(* Logix 5000 project; controller PLC_MCC1201_220AP1 vendor 1 type 14 code 164 rev 35.11; software revision 35.00; part 11 of 25 *)
(* tags used below, declared in another part *)
   AFI : ALIAS FOR B3[7].15;
   B175 : DINT[1];
   B176 : DINT[1];
   B180 : DINT[10];
   BT181_000 : MESSAGE;
   BT181_004 : MESSAGE;
   BT181_005 : MESSAGE;
   BT181_006 : MESSAGE;
   BT181_007 : MESSAGE;
   BT181_008 : MESSAGE;
   C183 : COUNTER[3];
   ConsumedFromCullet : UDT_CONSUMED_CULLET;
   ConsumedFromMCC1300 : UDT_CONSUMED_NEXT;
   CPU_FaultRecord : SYS_FaultRecord;
   CPU_LastFaultRecord : SYS_FaultRecord;
   From_Cullet : DINT[10];
   HMI_Always_ON : BOOL;   // HMI Always ON
   I : INT[128];
   M202_M1_DR : AXIS_CIP_DRIVE;
   M202_M1_DR_IN_MAJ : MOTION_INSTRUCTION;
   M202_M1_DR_IN_MAM : MOTION_INSTRUCTION;
   M202_M1_DR_IN_MAR : MOTION_INSTRUCTION;
   M202_M1_DR_IN_MAS : MOTION_INSTRUCTION;
   M202_M1_DR_IN_MCD : MOTION_INSTRUCTION;
   M202_M1_DR_IN_MRP : MOTION_INSTRUCTION;
   M202_M1_DR_OUT_MAJ : MOTION_INSTRUCTION;
   M202_M1_DR_OUT_MAM : MOTION_INSTRUCTION;
   M202_M1_DR_OUT_MAR : MOTION_INSTRUCTION;
   M202_M1_DR_OUT_MAS : MOTION_INSTRUCTION;
   M202_M1_DR_OUT_MCD : MOTION_INSTRUCTION;
   M202_M1_DR_OUT_MRP : MOTION_INSTRUCTION;
   M203_M1_DR : AXIS_CIP_DRIVE;
   M203_M1_DR_IN_MAJ : MOTION_INSTRUCTION;
   M203_M1_DR_IN_MAM : MOTION_INSTRUCTION;
   M203_M1_DR_IN_MAR : MOTION_INSTRUCTION;
   M203_M1_DR_IN_MAS : MOTION_INSTRUCTION;
   M203_M1_DR_IN_MCD : MOTION_INSTRUCTION;
   M203_M1_DR_IN_MRP : MOTION_INSTRUCTION;
   M203_M1_DR_OUT_MAJ : MOTION_INSTRUCTION;
   M203_M1_DR_OUT_MAM : MOTION_INSTRUCTION;
   M203_M1_DR_OUT_MAR : MOTION_INSTRUCTION;
   M203_M1_DR_OUT_MAS : MOTION_INSTRUCTION;
   M203_M1_DR_OUT_MCD : MOTION_INSTRUCTION;
   M203_M1_DR_OUT_MRP : MOTION_INSTRUCTION;
   M203DROP : MAC_DROPCONV;
   M204_M1_DR : AXIS_CIP_DRIVE;
   M204_M1_DR_IN_MAJ : MOTION_INSTRUCTION;
   M204_M1_DR_IN_MAM : MOTION_INSTRUCTION;
   M204_M1_DR_IN_MAR : MOTION_INSTRUCTION;
   M204_M1_DR_IN_MAS : MOTION_INSTRUCTION;
   M204_M1_DR_IN_MCD : MOTION_INSTRUCTION;
   M204_M1_DR_IN_MRP : MOTION_INSTRUCTION;
   M204_M1_DR_OUT_MAJ : MOTION_INSTRUCTION;
   M204_M1_DR_OUT_MAM : MOTION_INSTRUCTION;
   M204_M1_DR_OUT_MAR : MOTION_INSTRUCTION;
   M204_M1_DR_OUT_MAS : MOTION_INSTRUCTION;
   M204_M1_DR_OUT_MCD : MOTION_INSTRUCTION;
   M204_M1_DR_OUT_MRP : MOTION_INSTRUCTION;
   M205BREAKER : MAC_BREAKER;
   M206_M1_DR : AXIS_CIP_DRIVE;
   M206_M1_DR_IN_MAJ : MOTION_INSTRUCTION;
   M206_M1_DR_IN_MAM : MOTION_INSTRUCTION;
   M206_M1_DR_IN_MAR : MOTION_INSTRUCTION;
   M206_M1_DR_IN_MAS : MOTION_INSTRUCTION;
   M206_M1_DR_IN_MCD : MOTION_INSTRUCTION;
   M206_M1_DR_IN_MRP : MOTION_INSTRUCTION;
   M206_M1_DR_OUT_MAJ : MOTION_INSTRUCTION;
   M206_M1_DR_OUT_MAM : MOTION_INSTRUCTION;
   M206_M1_DR_OUT_MAR : MOTION_INSTRUCTION;
   M206_M1_DR_OUT_MAS : MOTION_INSTRUCTION;
   M206_M1_DR_OUT_MCD : MOTION_INSTRUCTION;
   M206_M1_DR_OUT_MRP : MOTION_INSTRUCTION;
   M207_M1_DR : AXIS_CIP_DRIVE;
   M207_M1_DR_IN_MAJ : MOTION_INSTRUCTION;
   M207_M1_DR_IN_MAM : MOTION_INSTRUCTION;
   M207_M1_DR_IN_MAR : MOTION_INSTRUCTION;
   M207_M1_DR_IN_MAS : MOTION_INSTRUCTION;
   M207_M1_DR_IN_MCD : MOTION_INSTRUCTION;
   M207_M1_DR_IN_MRP : MOTION_INSTRUCTION;
   M207_M1_DR_OUT_MAJ : MOTION_INSTRUCTION;
   M207_M1_DR_OUT_MAM : MOTION_INSTRUCTION;
   M207_M1_DR_OUT_MAR : MOTION_INSTRUCTION;
   M207_M1_DR_OUT_MAS : MOTION_INSTRUCTION;
   M207_M1_DR_OUT_MCD : MOTION_INSTRUCTION;
   M207_M1_DR_OUT_MRP : MOTION_INSTRUCTION;
   M208_M1_DR : AXIS_CIP_DRIVE;
   M208_M1_DR_IN_MAJ : MOTION_INSTRUCTION;
   M208_M1_DR_IN_MAM : MOTION_INSTRUCTION;
   M208_M1_DR_IN_MAR : MOTION_INSTRUCTION;
   M208_M1_DR_IN_MAS : MOTION_INSTRUCTION;
   M208_M1_DR_IN_MCD : MOTION_INSTRUCTION;
   M208_M1_DR_IN_MRP : MOTION_INSTRUCTION;
   M208_M1_DR_OUT_MAJ : MOTION_INSTRUCTION;
   M208_M1_DR_OUT_MAM : MOTION_INSTRUCTION;
   M208_M1_DR_OUT_MAR : MOTION_INSTRUCTION;
   M208_M1_DR_OUT_MAS : MOTION_INSTRUCTION;
   M208_M1_DR_OUT_MCD : MOTION_INSTRUCTION;
   M208_M1_DR_OUT_MRP : MOTION_INSTRUCTION;
   M209_M1_DR : AXIS_CIP_DRIVE;
   M209_M1_DR_IN_MAJ : MOTION_INSTRUCTION;
   M209_M1_DR_IN_MAM : MOTION_INSTRUCTION;
   M209_M1_DR_IN_MAR : MOTION_INSTRUCTION;
   M209_M1_DR_IN_MAS : MOTION_INSTRUCTION;
   M209_M1_DR_IN_MCD : MOTION_INSTRUCTION;
   M209_M1_DR_IN_MRP : MOTION_INSTRUCTION;
   M209_M1_DR_OUT_MAJ : MOTION_INSTRUCTION;
   M209_M1_DR_OUT_MAM : MOTION_INSTRUCTION;
   M209_M1_DR_OUT_MAR : MOTION_INSTRUCTION;
   M209_M1_DR_OUT_MAS : MOTION_INSTRUCTION;
   M209_M1_DR_OUT_MCD : MOTION_INSTRUCTION;
   M209_M1_DR_OUT_MRP : MOTION_INSTRUCTION;
   M210_M1_DR : AXIS_CIP_DRIVE;
   M210_M1_DR_IN_MAJ : MOTION_INSTRUCTION;
   M210_M1_DR_IN_MAM : MOTION_INSTRUCTION;
   M210_M1_DR_IN_MAR : MOTION_INSTRUCTION;
   M210_M1_DR_IN_MAS : MOTION_INSTRUCTION;
   M210_M1_DR_IN_MCD : MOTION_INSTRUCTION;
   M210_M1_DR_IN_MRP : MOTION_INSTRUCTION;
   M210_M1_DR_OUT_MAJ : MOTION_INSTRUCTION;
   M210_M1_DR_OUT_MAM : MOTION_INSTRUCTION;
   M210_M1_DR_OUT_MAR : MOTION_INSTRUCTION;
   M210_M1_DR_OUT_MAS : MOTION_INSTRUCTION;
   M210_M1_DR_OUT_MCD : MOTION_INSTRUCTION;
   M210_M1_DR_OUT_MRP : MOTION_INSTRUCTION;
   M211_M1_DR : AXIS_CIP_DRIVE;
   M211_M1_DR_IN_MAJ : MOTION_INSTRUCTION;
   M211_M1_DR_IN_MAM : MOTION_INSTRUCTION;
   M211_M1_DR_IN_MAR : MOTION_INSTRUCTION;
   M211_M1_DR_IN_MAS : MOTION_INSTRUCTION;
   M211_M1_DR_IN_MCD : MOTION_INSTRUCTION;
   M211_M1_DR_IN_MRP : MOTION_INSTRUCTION;
   M211_M1_DR_OUT_MAJ : MOTION_INSTRUCTION;
   M211_M1_DR_OUT_MAM : MOTION_INSTRUCTION;
   M211_M1_DR_OUT_MAR : MOTION_INSTRUCTION;
   M211_M1_DR_OUT_MAS : MOTION_INSTRUCTION;
   M211_M1_DR_OUT_MCD : MOTION_INSTRUCTION;
   M211_M1_DR_OUT_MRP : MOTION_INSTRUCTION;
   M212_M1_DR : AXIS_CIP_DRIVE;
   M212_M1_DR_IN_MAJ : MOTION_INSTRUCTION;
   M212_M1_DR_IN_MAM : MOTION_INSTRUCTION;
   M212_M1_DR_IN_MAR : MOTION_INSTRUCTION;
   M212_M1_DR_IN_MAS : MOTION_INSTRUCTION;
   M212_M1_DR_IN_MCD : MOTION_INSTRUCTION;
   M212_M1_DR_IN_MRP : MOTION_INSTRUCTION;
   M212_M1_DR_OUT_MAJ : MOTION_INSTRUCTION;
   M212_M1_DR_OUT_MAM : MOTION_INSTRUCTION;
   M212_M1_DR_OUT_MAR : MOTION_INSTRUCTION;
   M212_M1_DR_OUT_MAS : MOTION_INSTRUCTION;
   M212_M1_DR_OUT_MCD : MOTION_INSTRUCTION;
   M212_M1_DR_OUT_MRP : MOTION_INSTRUCTION;
   M213_M1_DR : AXIS_CIP_DRIVE;
   M213_M1_DR_IN_MAJ : MOTION_INSTRUCTION;
   M213_M1_DR_IN_MAM : MOTION_INSTRUCTION;
   M213_M1_DR_IN_MAR : MOTION_INSTRUCTION;
   M213_M1_DR_IN_MAS : MOTION_INSTRUCTION;
   M213_M1_DR_IN_MCD : MOTION_INSTRUCTION;
   M213_M1_DR_IN_MRP : MOTION_INSTRUCTION;
   M213_M1_DR_OUT_MAJ : MOTION_INSTRUCTION;
   M213_M1_DR_OUT_MAM : MOTION_INSTRUCTION;
   M213_M1_DR_OUT_MAR : MOTION_INSTRUCTION;
   M213_M1_DR_OUT_MAS : MOTION_INSTRUCTION;
   M213_M1_DR_OUT_MCD : MOTION_INSTRUCTION;
   M213_M1_DR_OUT_MRP : MOTION_INSTRUCTION;
   M213A_M1_DR_IN_MAJ : MOTION_INSTRUCTION;
   M213A_M1_DR_IN_MAM : MOTION_INSTRUCTION;
   M213A_M1_DR_IN_MAR : MOTION_INSTRUCTION;
   M213A_M1_DR_IN_MAS : MOTION_INSTRUCTION;
   M213A_M1_DR_IN_MCD : MOTION_INSTRUCTION;
   M213A_M1_DR_IN_MRP : MOTION_INSTRUCTION;
   M213A_M1_DR_OUT_MAJ : MOTION_INSTRUCTION;
   M213A_M1_DR_OUT_MAM : MOTION_INSTRUCTION;
   M213A_M1_DR_OUT_MAR : MOTION_INSTRUCTION;
   M213A_M1_DR_OUT_MAS : MOTION_INSTRUCTION;
   M213A_M1_DR_OUT_MCD : MOTION_INSTRUCTION;
   M213A_M1_DR_OUT_MRP : MOTION_INSTRUCTION;
   M213B_M1_DR_IN_MAJ : MOTION_INSTRUCTION;
   M213B_M1_DR_IN_MAM : MOTION_INSTRUCTION;
   M213B_M1_DR_IN_MAR : MOTION_INSTRUCTION;
   M213B_M1_DR_IN_MAS : MOTION_INSTRUCTION;
   M213B_M1_DR_IN_MCD : MOTION_INSTRUCTION;
   M213B_M1_DR_IN_MRP : MOTION_INSTRUCTION;
   M213B_M1_DR_OUT_MAJ : MOTION_INSTRUCTION;
   M213B_M1_DR_OUT_MAM : MOTION_INSTRUCTION;
   M213B_M1_DR_OUT_MAR : MOTION_INSTRUCTION;
   M213B_M1_DR_OUT_MAS : MOTION_INSTRUCTION;
   M213B_M1_DR_OUT_MCD : MOTION_INSTRUCTION;
   M213B_M1_DR_OUT_MRP : MOTION_INSTRUCTION;
   M214_M1_DR : AXIS_CIP_DRIVE;
   M214_M1_DR_IN_MAJ : MOTION_INSTRUCTION;
   M214_M1_DR_IN_MAM : MOTION_INSTRUCTION;
   M214_M1_DR_IN_MAR : MOTION_INSTRUCTION;
   M214_M1_DR_IN_MAS : MOTION_INSTRUCTION;
   M214_M1_DR_IN_MCD : MOTION_INSTRUCTION;
   M214_M1_DR_IN_MRP : MOTION_INSTRUCTION;
   M214_M1_DR_OUT_MAJ : MOTION_INSTRUCTION;
   M214_M1_DR_OUT_MAM : MOTION_INSTRUCTION;
   M214_M1_DR_OUT_MAR : MOTION_INSTRUCTION;
   M214_M1_DR_OUT_MAS : MOTION_INSTRUCTION;
   M214_M1_DR_OUT_MCD : MOTION_INSTRUCTION;
   M214_M1_DR_OUT_MRP : MOTION_INSTRUCTION;
   M215_M1_DR : AXIS_CIP_DRIVE;
   M215_M1_DR_IN_MAJ : MOTION_INSTRUCTION;
   M215_M1_DR_IN_MAM : MOTION_INSTRUCTION;
   M215_M1_DR_IN_MAR : MOTION_INSTRUCTION;
   M215_M1_DR_IN_MAS : MOTION_INSTRUCTION;
   M215_M1_DR_IN_MCD : MOTION_INSTRUCTION;
   M215_M1_DR_IN_MRP : MOTION_INSTRUCTION;
   M215_M1_DR_OUT_MAJ : MOTION_INSTRUCTION;
   M215_M1_DR_OUT_MAM : MOTION_INSTRUCTION;
   M215_M1_DR_OUT_MAR : MOTION_INSTRUCTION;
   M215_M1_DR_OUT_MAS : MOTION_INSTRUCTION;
   M215_M1_DR_OUT_MCD : MOTION_INSTRUCTION;
   M215_M1_DR_OUT_MRP : MOTION_INSTRUCTION;
   M216_M1_DR : AXIS_CIP_DRIVE;
   M216_M1_DR_IN_MAJ : MOTION_INSTRUCTION;
   M216_M1_DR_IN_MAM : MOTION_INSTRUCTION;
   M216_M1_DR_IN_MAR : MOTION_INSTRUCTION;
   M216_M1_DR_IN_MAS : MOTION_INSTRUCTION;
   M216_M1_DR_IN_MCD : MOTION_INSTRUCTION;
   M216_M1_DR_IN_MRP : MOTION_INSTRUCTION;
   M216_M1_DR_OUT_MAJ : MOTION_INSTRUCTION;
   M216_M1_DR_OUT_MAM : MOTION_INSTRUCTION;
   M216_M1_DR_OUT_MAR : MOTION_INSTRUCTION;
   M216_M1_DR_OUT_MAS : MOTION_INSTRUCTION;
   M216_M1_DR_OUT_MCD : MOTION_INSTRUCTION;
   M216_M1_DR_OUT_MRP : MOTION_INSTRUCTION;
   M217_M1_DR : AXIS_CIP_DRIVE;
   M217_M1_DR_IN_MAJ : MOTION_INSTRUCTION;
   M217_M1_DR_IN_MAM : MOTION_INSTRUCTION;
   M217_M1_DR_IN_MAR : MOTION_INSTRUCTION;
   M217_M1_DR_IN_MAS : MOTION_INSTRUCTION;
   M217_M1_DR_IN_MCD : MOTION_INSTRUCTION;
   M217_M1_DR_IN_MRP : MOTION_INSTRUCTION;
   M217_M1_DR_OUT_MAJ : MOTION_INSTRUCTION;
   M217_M1_DR_OUT_MAM : MOTION_INSTRUCTION;
   M217_M1_DR_OUT_MAR : MOTION_INSTRUCTION;
   M217_M1_DR_OUT_MAS : MOTION_INSTRUCTION;
   M217_M1_DR_OUT_MCD : MOTION_INSTRUCTION;
   M217_M1_DR_OUT_MRP : MOTION_INSTRUCTION;
   M218_M1_DR : AXIS_CIP_DRIVE;
   M218_M1_DR_IN_MAJ : MOTION_INSTRUCTION;
   M218_M1_DR_IN_MAM : MOTION_INSTRUCTION;
   M218_M1_DR_IN_MAR : MOTION_INSTRUCTION;
   M218_M1_DR_IN_MAS : MOTION_INSTRUCTION;
   M218_M1_DR_IN_MCD : MOTION_INSTRUCTION;
   M218_M1_DR_IN_MRP : MOTION_INSTRUCTION;
   M218_M1_DR_OUT_MAJ : MOTION_INSTRUCTION;
   M218_M1_DR_OUT_MAM : MOTION_INSTRUCTION;
   M218_M1_DR_OUT_MAR : MOTION_INSTRUCTION;
   M218_M1_DR_OUT_MAS : MOTION_INSTRUCTION;
(* CommandLogic, continued *)

ROUTINE Main   (* ladder *)
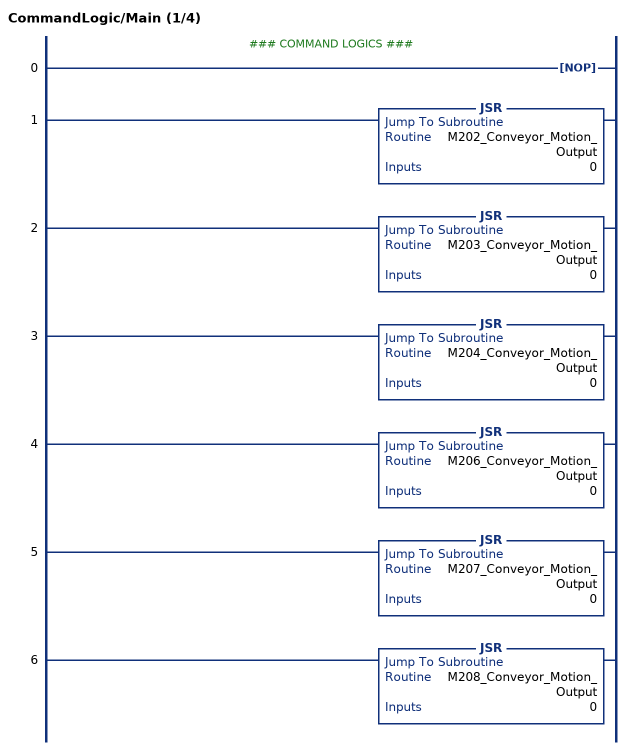
   // ### COMMAND LOGICS ###
   0: NOP();
   1: JSR(M202_Conveyor_Motion_Output,0);
   2: JSR(M203_Conveyor_Motion_Output,0);
   3: JSR(M204_Conveyor_Motion_Output,0);
   4: JSR(M206_Conveyor_Motion_Output,0);
   5: JSR(M207_Conveyor_Motion_Output,0);
   6: JSR(M208_Conveyor_Motion_Output,0);
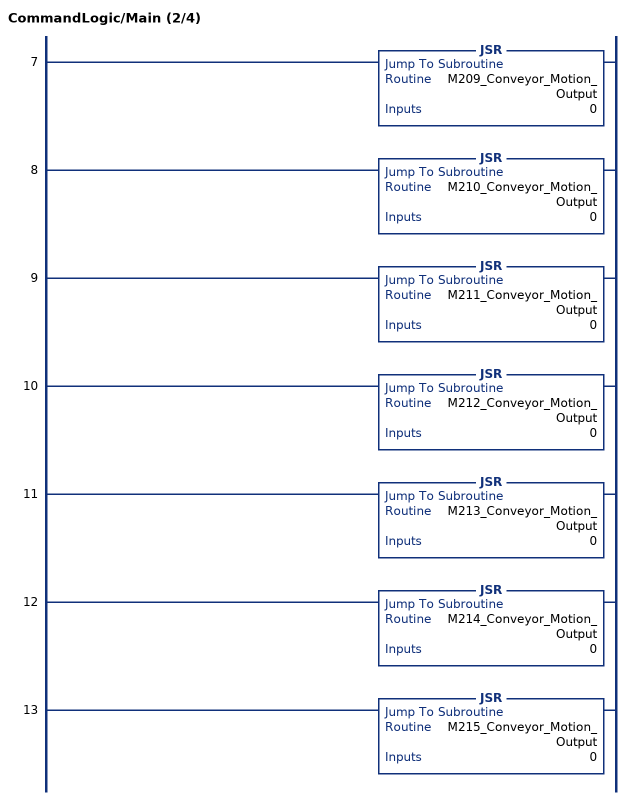
   7: JSR(M209_Conveyor_Motion_Output,0);
   8: JSR(M210_Conveyor_Motion_Output,0);
   9: JSR(M211_Conveyor_Motion_Output,0);
   10: JSR(M212_Conveyor_Motion_Output,0);
   11: JSR(M213_Conveyor_Motion_Output,0);
   12: JSR(M214_Conveyor_Motion_Output,0);
   13: JSR(M215_Conveyor_Motion_Output,0);
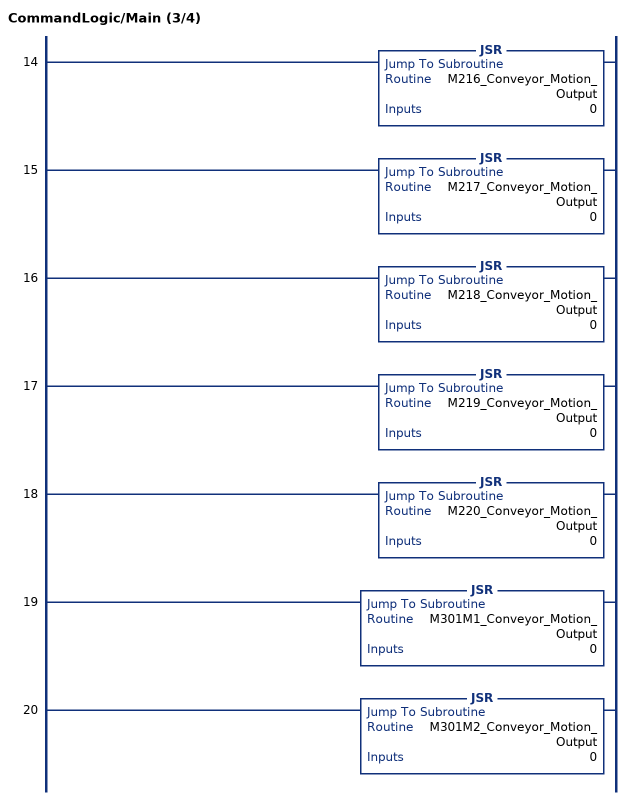
   14: JSR(M216_Conveyor_Motion_Output,0);
   15: JSR(M217_Conveyor_Motion_Output,0);
   16: JSR(M218_Conveyor_Motion_Output,0);
   17: JSR(M219_Conveyor_Motion_Output,0);
   18: JSR(M220_Conveyor_Motion_Output,0);
   19: JSR(M301M1_Conveyor_Motion_Output,0);
   20: JSR(M301M2_Conveyor_Motion_Output,0);
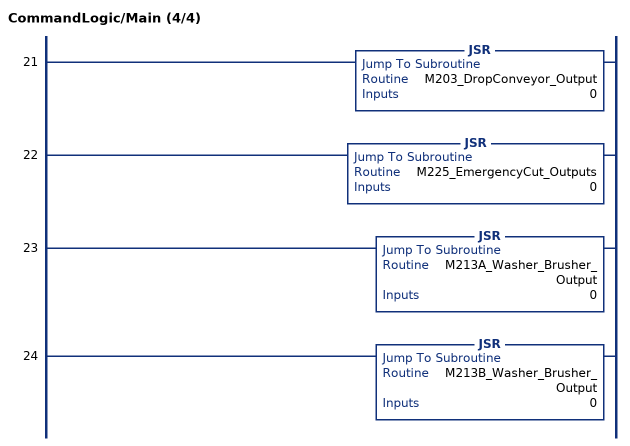
   21: JSR(M203_DropConveyor_Output,0);
   22: JSR(M225_EmergencyCut_Outputs,0);
   23: JSR(M213A_Washer_Brusher_Output,0);
   24: JSR(M213B_Washer_Brusher_Output,0);
END_ROUTINE
END_PROGRAM

PROGRAM ControllerErrors   (* main routine Main *)

ROUTINE Main   (* ladder *)
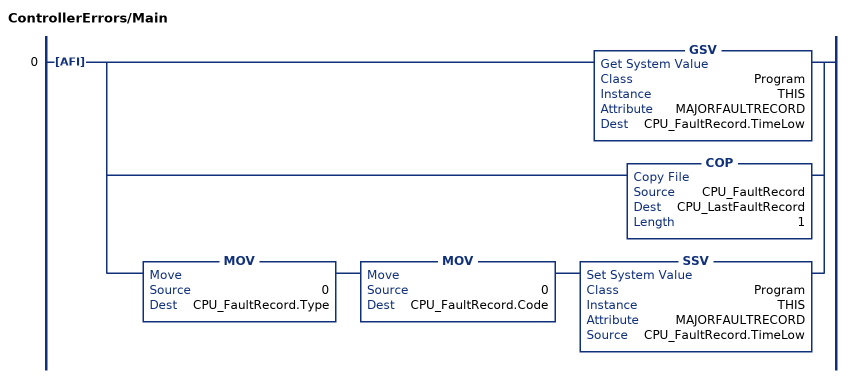
   0: AFI()[GSV(Program,THIS,MAJORFAULTRECORD,CPU_FaultRecord.TimeLow) ,COP(CPU_FaultRecord,CPU_LastFaultRecord,1) ,MOV(0,CPU_FaultRecord.Type) MOV(0,CPU_FaultRecord.Code) SSV(Program,THIS,MAJORFAULTRECORD,CPU_FaultRecord.TimeLow) ];
END_ROUTINE
END_PROGRAM

PROGRAM MainProgram   (* main routine MainRoutine *)
VAR
   dMaxLehrSpeed : DINT := 20000;
   dMinLehrSpeed : DINT := 1270;
   GP_M225_AccessArea_FarSide : GP_AccessArea := (IN_xConditionOkForcedAccess := 1);
   GP_M225_AccessArea_FarSide_STC : GP_AccessArea_STC := (OSR_xAccessRequest := 1, OSR_xAccessAcceptedAndButtonReleased := 1, OSR_xRemoveAccess := 1, OSR_xRemoveAccessNotAccepted := 1);
   GP_M225_AccessArea_OpSide : GP_AccessArea := (IN_xConditionOkForcedAccess := 1);
   GP_M225_AccessArea_OpSide_STC : GP_AccessArea_STC := (OSR_xAccessRequest := 1, OSR_xAccessAcceptedAndButtonReleased := 1, OSR_xRemoveAccess := 1, OSR_xRemoveAccessNotAccepted := 1);
   GP_RibbonTracking_GetRibbonData : GP_RibbonTracking_GetRibbonData;
   GP_RibbonTracking_UpdateGlassBreak : GP_RibbonTracking_UpdateGlassBreak;
   LEHR_dActualSpeedValue_mm_min : DINT;
   LEHR_dActualSpeedValueToConveyor_mm_min : DINT;
   LEHR_dLehrPositionAdvancement : DINT;
   SnaprollHMW_dOffset_cmm : DINT;
   SnaprollUPS_DistanceFromSnaproll_cmm : DINT := 4663000;
   SnaprollUPS_xOS_NewCut : BOOL;
   SnaprollUPS_xOSR : BOOL;
   SnaprollUPS_xOutputRise : BOOL;
   tmOF_retainSnaprolUPS : TIMER;
   TMP_dDistanceBetweenCut : DINT := 273986272;
   TMP_dDummy : DINT := 4215000;
   TMP_dEncoderCutPosition : DINT;
   TMP_dSnaprollCut_cmm : DINT := 4663000;
   TMP_dValue : DINT;
   TMP_xCutOnSnaproll_cmm : BOOL;
   TMP_xDummy : BOOL;
   TMP_xSimulationMode : BOOL;
   xAlwaysOFF : BOOL;
   xAlwaysON : BOOL := 1;
   xDebugOFF : BOOL;
END_VAR

ROUTINE _010_Input_Mapping   (* structured text *)
   
   //Always ON bit for HMI
   HMI_Always_ON := 1;
   
   //INPUT
   
   //Z200 UPS ZONE (UNTIL MAIN CRUSHER)
   Z200_UPS.INPUT_x24vdcVoltageOn := A152AP1:1:I.Pt00.Data;
   Z200_UPS.INPUT_xUPSEmergencyON := A152AP1:1:I.Pt04.Data;
   Z200_UPS.INPUT_xEmLocUps1 := A152AP1:6:I.Pt11.Data; //A33SB2 UPS Emergency Button M203DROP OPERATOR SIDE
   Z200_UPS.INPUT_xEmLocUps2 := A152AP1:6:I.Pt14.Data; //A33SB3 UPS Emergency Button M203DROP FAR SIDE
   Z200_UPS.INPUT_xEmLocUps3 := A152AP1:8:I.Pt02.Data; //A33SB4 UPS Emergency Button M225
   Z200_UPS.INPUT_xEmLocUps4 := A152AP1:8:I.Pt07.Data; //A33SB5 UPS Emergency Button CS4225
   
   //Z200 UNDER CUTTING TRANSPORT ZONE
   
   Z200.INPUT_x24VdcVoltageON := A152AP1:1:I.Pt00.Data;
   //spare
   Z200.INPUT_xEmergencyLocalization1 := A152AP1:1:I.Pt02.Data;//A33SB1 Main Emergency Button MCC1201
   //spare
   Z200.INPUT_xUPSEmergencyON := A152AP1:1:I.Pt04.Data;
   Z200.INPUT_xMainEmergencyON := A152AP1:1:I.Pt05.Data;
   //spare
   Z200.INPUT_xMainSwitch := A152AP1:1:I.Pt07.Data;
   Z200.INPUT_xPowerFailure120V_Auxiliary1 := A152AP1:1:I.Pt08.Data;
   Z200.INPUT_xPowerFailure120V_Auxiliary2 := A152AP1:1:I.Pt09.Data;
   Z200.INPUT_xPowerSupplyOK := A152AP1:1:I.Pt10.Data;
   Z200.INPUT_xPowerSupply24VLogic1 := A152AP1:1:I.Pt11.Data;
   Z200.INPUT_xPowerSupply24VLogic2 := A152AP1:1:I.Pt12.Data;
   Z200.INPUT_xPowerSupply24VLogic3 := A152AP1:1:I.Pt13.Data;
   Z200.INPUT_xPowerSupply24VLogic4 := A152AP1:1:I.Pt14.Data;
   Z200.INPUT_xEthernetSwitchFault := A152AP1:1:I.Pt15.Data;
   
   Z200.INPUT_xProtectionPowerSupplyConditioner1 := A152AP1:2:I.Pt15.Data;
   Z200.INPUT_xProtectionPowerSupplyConditioner2 := A152AP1:4:I.Pt15.Data;
   
   Z200.INPUT_xEmergencyLocalization2 := A152AP1:7:I.Pt00.Data; //A34SB1 Main Emergency Button M203DROP OPERATOR SIDE
   Z200.INPUT_xEmergencyLocalization3 := A152AP1:7:I.Pt01.Data; //A34SB2 Main Emergency Button M203DROP FAR SIDE
   
   Z200.INPUT_xAlarmSilence := A152AP1:11:I.Pt08.Data;
   Z200.INPUT_xAlarmReset := A152AP1:11:I.Pt09.Data;
   
   
   //M202
   M2xx_CONVEYOR[0].INPUT_xProtectionRot := A152AP1:2:I.Pt00.Data;
   M2xx_CONVEYOR[0].INPUT_xProtectionFan := A152AP1:2:I.Pt01.Data;
   M2xx_CONVEYOR[0].INPUT_xLocalSafetySwitch := A152AP1:6:I.Pt00.Data;
   M2xx_CONVEYOR[0].INPUT_xThermalProbe := A152AP1:6:I.Pt01.Data;
   M2xx_CONVEYOR[0].INPUT_xDriveInhibit := M202_M1_DR.CIPAxisState = 9;
   M2xx_CONVEYOR[0].INPUT_xDriveReady := M202_M1_DR.ServoActionStatus;
   M2xx_CONVEYOR[0].INPUT_xDriveError := M202_M1_DR.AxisFault <> 0 OR M202_M1_DR.ModuleFaults <> 0;
   M2xx_CONVEYOR[0].INPUT_xRotationFeedback := M202_M1_DR.MotionStatus <> 0;
   
   //M203
   M2xx_CONVEYOR[1].INPUT_xProtectionRot := A152AP1:2:I.Pt02.Data;
   M2xx_CONVEYOR[1].INPUT_xProtectionFan := A152AP1:2:I.Pt03.Data;
   M2xx_CONVEYOR[1].INPUT_xLocalSafetySwitch := A152AP1:6:I.Pt03.Data;
   M2xx_CONVEYOR[1].INPUT_xThermalProbe := A152AP1:6:I.Pt04.Data;
   M2xx_CONVEYOR[1].INPUT_xDriveInhibit := M203_M1_DR.CIPAxisState = 9;
   M2xx_CONVEYOR[1].INPUT_xDriveReady := M203_M1_DR.ServoActionStatus;
   M2xx_CONVEYOR[1].INPUT_xDriveError := M203_M1_DR.AxisFault <> 0 OR M203_M1_DR.ModuleFaults <> 0;
   M2xx_CONVEYOR[1].INPUT_xRotationFeedback := M203_M1_DR.MotionStatus <> 0;
   
   //M203DROP
   M203DROP.INPUT_xUpPosition := A152AP1:6:I.Pt05.Data;
   M203DROP.INPUT_xDownPosition := A152AP1:6:I.Pt06.Data;
   M203DROP.INPUT_xTiltingSafetyBarDisinsered := A152AP1:6:I.Pt07.Data;
   M203DROP.INPUT_xDoorOpenTiltingAreaOpSide := A152AP1:6:I.Pt09.Data;
   M203DROP.INPUT_xUpDownPushbuttonOpSide := A152AP1:6:I.Pt10.Data;
   M203DROP.INPUT_xDoorOpenTiltingAreaOpSide := A152AP1:6:I.Pt12.Data;
   M203DROP.INPUT_xUpDownPushbuttonOpSide := A152AP1:6:I.Pt13.Data;
   
   //M204
   M2xx_CONVEYOR[2].INPUT_xProtectionRot := A152AP1:2:I.Pt04.Data;
   M2xx_CONVEYOR[2].INPUT_xProtectionFan := xAlwaysON;
   M2xx_CONVEYOR[2].INPUT_xLocalSafetySwitch := A152AP1:7:I.Pt03.Data;
   M2xx_CONVEYOR[2].INPUT_xThermalProbe := A152AP1:7:I.Pt04.Data;
   M2xx_CONVEYOR[2].INPUT_xDriveInhibit := M204_M1_DR.CIPAxisState = 9;
   M2xx_CONVEYOR[2].INPUT_xDriveReady := M204_M1_DR.ServoActionStatus;
   M2xx_CONVEYOR[2].INPUT_xDriveError := M204_M1_DR.AxisFault <> 0 OR M204_M1_DR.ModuleFaults <> 0;
   M2xx_CONVEYOR[2].INPUT_xRotationFeedback := M204_M1_DR.MotionStatus <> 0;
   
   //M205 BREAKER
   M205BREAKER.INPUT_xProtectionBreaker := A152AP1:2:I.Pt06.Data;
   M205BREAKER.INPUT_xFeedBackBreakerRotation := A152AP1:2:I.Pt07.Data;
   M205BREAKER.INPUT_xFeedbackExclusionInductance := A152AP1:2:I.Pt08.Data;
   M205BREAKER.INPUT_xLocalSafetySwitch := A152AP1:7:I.Pt05.Data;
   M205BREAKER.INPUT_xBreakerControlRotation := A152AP1:7:I.Pt06.Data;
   
   //M225 EMERGENCY XCUT
   M225.INPUT_xProtectionTraslation := A152AP1:2:I.Pt09.Data;
   M225.INPUT_xProtectionFan := A152AP1:2:I.Pt10.Data;
   M225.INPUT_xAreaSafety := A152AP1:2:I.Pt11.Data;
   M225.INPUT_xLocalSafetySwitch := A152AP1:7:I.Pt08.Data;
   M225.INPUT_xThermalProbe := A152AP1:7:I.Pt09.Data;
   M225.INPUT_xHomePosition := A152AP1:7:I.Pt10.Data;
   M225.INPUT_xOverstrokeFW := A152AP1:7:I.Pt11.Data;
   M225.INPUT_xOverstrokeBW := A152AP1:7:I.Pt12.Data;
   M225.INPUT_xCompressedAirPresence := A152AP1:7:I.Pt13.Data;
   M225.INPUT_xLubricationTest := A152AP1:7:I.Pt14.Data;
   M225.INPUT_xCuttingHeadTest := A152AP1:7:I.Pt15.Data;
   M225.INPUT_xCuttingHeadHigh := A152AP1:8:I.Pt00.Data;
   M225.INPUT_xCuttingSafety := A152AP1:8:I.Pt01.Data; //photocell sensor
   M225.INPUT_xOpeningDoorLocalizationFarSide := A152AP1:8:I.Pt03.Data;
   M225.INPUT_xResetAreaSafetiesFarSide := A152AP1:8:I.Pt04.Data;
   M225.INPUT_xAccessAreaRequestFarSide := A152AP1:8:I.Pt05.Data;
   
   //CS4225 EMERGENCY XCUT CONSOLLE
   M225.INPUT_xOpeningDoorLocalizationOpSide := A152AP1:8:I.Pt06.Data;
   M225.INPUT_xResetAreaSafetiesOpSide := A152AP1:8:I.Pt08.Data;
   M225.INPUT_xAccessAreaRequestOpSide := A152AP1:8:I.Pt09.Data;
   M225.INPUT_xManual := A152AP1:8:I.Pt10.Data;
   M225.INPUT_xAutomatic := A152AP1:8:I.Pt11.Data;
   M225.INPUT_xAlarmOff := A152AP1:8:I.Pt12.Data;
   M225.INPUT_xCutInterruption := A152AP1:8:I.Pt13.Data;
   M225.INPUT_xStartCut := A152AP1:8:I.Pt14.Data;
   M225.INPUT_xStopCut := A152AP1:8:I.Pt15.Data;
   
   //M206
   M2xx_CONVEYOR[3].INPUT_xProtectionRot := A152AP1:3:I.Pt00.Data;
   M2xx_CONVEYOR[3].INPUT_xProtectionFan := xAlwaysON;
   M2xx_CONVEYOR[3].INPUT_xLocalSafetySwitch := A152AP1:9:I.Pt00.Data;
   M2xx_CONVEYOR[3].INPUT_xThermalProbe := A152AP1:9:I.Pt01.Data;
   M2xx_CONVEYOR[3].INPUT_xDriveInhibit := M206_M1_DR.CIPAxisState = 9;
   M2xx_CONVEYOR[3].INPUT_xDriveReady := M206_M1_DR.ServoActionStatus;
   M2xx_CONVEYOR[3].INPUT_xDriveError := M206_M1_DR.AxisFault <> 0 OR M206_M1_DR.ModuleFaults <> 0;
   M2xx_CONVEYOR[3].INPUT_xRotationFeedback := M206_M1_DR.MotionStatus <> 0;
   
   //M207
   M2xx_CONVEYOR[4].INPUT_xProtectionRot := A152AP1:3:I.Pt01.Data;
   M2xx_CONVEYOR[4].INPUT_xProtectionFan := xAlwaysON;
   M2xx_CONVEYOR[4].INPUT_xLocalSafetySwitch := A152AP1:9:I.Pt02.Data;
   M2xx_CONVEYOR[4].INPUT_xThermalProbe := A152AP1:9:I.Pt03.Data;
   M2xx_CONVEYOR[4].INPUT_xDriveInhibit := M207_M1_DR.CIPAxisState = 9;
   M2xx_CONVEYOR[4].INPUT_xDriveReady := M207_M1_DR.ServoActionStatus;
   M2xx_CONVEYOR[4].INPUT_xDriveError := M207_M1_DR.AxisFault <> 0 OR M207_M1_DR.ModuleFaults <> 0;
   M2xx_CONVEYOR[4].INPUT_xRotationFeedback := M207_M1_DR.MotionStatus <> 0;
   
   //M208
   M2xx_CONVEYOR[5].INPUT_xProtectionRot := A152AP1:3:I.Pt02.Data;
   M2xx_CONVEYOR[5].INPUT_xProtectionFan := xAlwaysON;
   M2xx_CONVEYOR[5].INPUT_xLocalSafetySwitch := A152AP1:9:I.Pt04.Data;
   M2xx_CONVEYOR[5].INPUT_xThermalProbe := A152AP1:9:I.Pt05.Data;
   M2xx_CONVEYOR[5].INPUT_xDriveInhibit := M208_M1_DR.CIPAxisState = 9;
   M2xx_CONVEYOR[5].INPUT_xDriveReady := M208_M1_DR.ServoActionStatus;
   M2xx_CONVEYOR[5].INPUT_xDriveError := M208_M1_DR.AxisFault <> 0 OR M208_M1_DR.ModuleFaults <> 0;
   M2xx_CONVEYOR[5].INPUT_xRotationFeedback := M208_M1_DR.MotionStatus <> 0;
   
   //M209
   M2xx_CONVEYOR[6].INPUT_xProtectionRot := A152AP1:3:I.Pt03.Data;
   M2xx_CONVEYOR[6].INPUT_xProtectionFan := xAlwaysON;
   M2xx_CONVEYOR[6].INPUT_xLocalSafetySwitch := A152AP1:9:I.Pt06.Data;
   M2xx_CONVEYOR[6].INPUT_xThermalProbe := A152AP1:9:I.Pt07.Data;
   M2xx_CONVEYOR[6].INPUT_xDriveInhibit := M209_M1_DR.CIPAxisState = 9;
   M2xx_CONVEYOR[6].INPUT_xDriveReady := M209_M1_DR.ServoActionStatus;
   M2xx_CONVEYOR[6].INPUT_xDriveError := M209_M1_DR.AxisFault <> 0 OR M209_M1_DR.ModuleFaults <> 0;
   M2xx_CONVEYOR[6].INPUT_xRotationFeedback := M209_M1_DR.MotionStatus <> 0;
   
   //M210
   M2xx_CONVEYOR[7].INPUT_xProtectionRot := A152AP1:3:I.Pt04.Data;
   M2xx_CONVEYOR[7].INPUT_xProtectionFan := xAlwaysON;
   M2xx_CONVEYOR[7].INPUT_xLocalSafetySwitch := A152AP1:9:I.Pt08.Data;
   M2xx_CONVEYOR[7].INPUT_xThermalProbe := A152AP1:9:I.Pt09.Data;
   M2xx_CONVEYOR[7].INPUT_xDriveInhibit := M210_M1_DR.CIPAxisState = 9;
   M2xx_CONVEYOR[7].INPUT_xDriveReady := M210_M1_DR.ServoActionStatus;
   M2xx_CONVEYOR[7].INPUT_xDriveError := M210_M1_DR.AxisFault <> 0 OR M210_M1_DR.ModuleFaults <> 0;
   M2xx_CONVEYOR[7].INPUT_xRotationFeedback := M210_M1_DR.MotionStatus <> 0;
   
   //M211
   M2xx_CONVEYOR[8].INPUT_xProtectionRot := A152AP1:3:I.Pt05.Data;
   M2xx_CONVEYOR[8].INPUT_xProtectionFan := xAlwaysON;
   M2xx_CONVEYOR[8].INPUT_xLocalSafetySwitch := A152AP1:9:I.Pt10.Data;
   M2xx_CONVEYOR[8].INPUT_xThermalProbe := A152AP1:9:I.Pt11.Data;
   M2xx_CONVEYOR[8].INPUT_xDriveInhibit := M211_M1_DR.CIPAxisState = 9;
   M2xx_CONVEYOR[8].INPUT_xDriveReady := M211_M1_DR.ServoActionStatus;
   M2xx_CONVEYOR[8].INPUT_xDriveError := M211_M1_DR.AxisFault <> 0 OR M211_M1_DR.ModuleFaults <> 0;
   M2xx_CONVEYOR[8].INPUT_xRotationFeedback := M211_M1_DR.MotionStatus <> 0;
   
   //M212
   M2xx_CONVEYOR[9].INPUT_xProtectionRot := A152AP1:3:I.Pt06.Data;
   M2xx_CONVEYOR[9].INPUT_xProtectionFan := xAlwaysON;
   M2xx_CONVEYOR[9].INPUT_xLocalSafetySwitch := A152AP1:9:I.Pt12.Data;
   M2xx_CONVEYOR[9].INPUT_xThermalProbe := A152AP1:9:I.Pt13.Data;
   M2xx_CONVEYOR[9].INPUT_xDriveInhibit := M212_M1_DR.CIPAxisState = 9;
   M2xx_CONVEYOR[9].INPUT_xDriveReady := M212_M1_DR.ServoActionStatus;
   M2xx_CONVEYOR[9].INPUT_xDriveError := M212_M1_DR.AxisFault <> 0 OR M212_M1_DR.ModuleFaults <> 0;
   M2xx_CONVEYOR[9].INPUT_xRotationFeedback := M212_M1_DR.MotionStatus <> 0;
   
   //M213
   M2xx_CONVEYOR[10].INPUT_xProtectionRot := A152AP1:3:I.Pt07.Data;
   M2xx_CONVEYOR[10].INPUT_xProtectionFan := xAlwaysON;
   M2xx_CONVEYOR[10].INPUT_xLocalSafetySwitch := A152AP1:9:I.Pt14.Data;
   M2xx_CONVEYOR[10].INPUT_xThermalProbe := A152AP1:9:I.Pt15.Data;
   M2xx_CONVEYOR[10].INPUT_xDriveInhibit := M213_M1_DR.CIPAxisState = 9;
   M2xx_CONVEYOR[10].INPUT_xDriveReady := M213_M1_DR.ServoActionStatus;
   M2xx_CONVEYOR[10].INPUT_xDriveError := M213_M1_DR.AxisFault <> 0 OR M213_M1_DR.ModuleFaults <> 0;
   M2xx_CONVEYOR[10].INPUT_xRotationFeedback := M213_M1_DR.MotionStatus <> 0;